(* Logix 5000 project; controller FV vendor 1 type 14 code 217 rev 31.11; software revision 31.00; part 39 of 63 *)
(* tags used below, declared in another part *)
   FV_FV10C : PlantItem;   // FV10C
   FV_FV10C_RawOutput : ALIAS FOR Remote_IO:2:O.Data.2;   // FV_FV10C FV 10 cone cooling valve
   FV_FV10J : PlantItem;   // FV10J
   FV_FV10J_RawOutput : ALIAS FOR Remote_IO:2:O.Data.3;   // FV_FV10J FV 10 jacket cooling valve
   FV_FV11C : PlantItem;   // FV11C
   FV_FV11C_RawOutput : ALIAS FOR Remote_IO:2:O.Data.4;   // FV_FV11C FV 11 cone cooling valve
   FV_FV11J : PlantItem;   // FV11J
   FV_FV11J_RawOutput : ALIAS FOR Remote_IO:2:O.Data.5;   // FV_FV11J FV 11 jacket cooling valve
   FV_FV12C : PlantItem;   // FV12C
   FV_FV12C_RawOutput : ALIAS FOR Remote_IO:2:O.Data.6;   // FV_FV12C FV 12 cone cooling valve
   FV_FV12J : PlantItem;   // FV12J
   FV_FV12J_RawOutput : ALIAS FOR Remote_IO:2:O.Data.7;   // FV_FV12J FV 12 jacket cooling valve
   FV_FV13C : PlantItem;   // FV13C
   FV_FV13C_RawOutput : ALIAS FOR Remote_IO:2:O.Data.8;   // FV_FV13C FV 13 cone cooling valve
   FV_FV13J : PlantItem;   // FV13J
   FV_FV13J_RawOutput : ALIAS FOR Remote_IO:2:O.Data.9;   // FV_FV13J FV 13 jacket cooling valve
   FV_FV14C : PlantItem;   // FV14C
   FV_FV14C_RawOutput : ALIAS FOR Remote_IO:2:O.Data.10;   // FV_FV14C FV 14 cone cooling valve
   FV_FV14J : PlantItem;   // FV14J
   FV_FV14J_RawOutput : ALIAS FOR Remote_IO:2:O.Data.11;   // FV_FV14J FV 14 jacket cooling valve
   FV_FV15C : PlantItem;   // FV15C
   FV_FV15C_RawOutput : ALIAS FOR Remote_IO:2:O.Data.12;   // FV_FV15C FV 15 cone cooling valve
   FV_FV15J : PlantItem;   // FV15J
   FV_FV15J_RawOutput : ALIAS FOR Remote_IO:2:O.Data.13;   // FV_FV15J FV 15 jacket cooling valve
   FV_FV16C : PlantItem;   // FV16C
   FV_FV16C_RawOutput : ALIAS FOR Remote_IO:2:O.Data.14;   // FV_FV16C FV 16 cone cooling valve
   FV_FV16J : PlantItem;   // FV16J
   FV_FV16J_RawOutput : ALIAS FOR Remote_IO:2:O.Data.15;   // FV_FV16J FV 16 jacket cooling valve
   FV_FV17C : PlantItem;   // FV17C
   FV_FV17C_RawOutput : ALIAS FOR Remote_IO:3:O.Data.0;   // FV_FV17C FV 17 cone cooling valve
   FV_FV17J : PlantItem;   // FV17J
   FV_FV17J_RawOutput : ALIAS FOR Remote_IO:3:O.Data.1;   // FV_FV17J FV 17 jacket cooling valve
   FV_FV18C : PlantItem;   // FV18C
   FV_FV18C_RawOutput : ALIAS FOR Remote_IO:3:O.Data.2;   // FV_FV18C FV 18 cone cooling valve
   FV_FV18J : PlantItem;   // FV18J
   FV_FV18J_RawOutput : ALIAS FOR Remote_IO:3:O.Data.3;   // FV_FV18J FV 18 jacket cooling valve
   FV_FV19C : PlantItem;   // FV19C
   FV_FV19C_RawOutput : ALIAS FOR Remote_IO:3:O.Data.4;   // FV_FV19C FV 19 cone cooling valve
   FV_FV19J : PlantItem;   // FV19J
   FV_FV19J_RawOutput : ALIAS FOR Remote_IO:3:O.Data.5;   // FV_FV19J FV 19 jacket cooling valve
   FV_FV1C : PlantItem;   // FV1C
   FV_FV1C_RawOutput : ALIAS FOR Remote_IO:1:O.Data.0;   // FV_FV1C FV 1 cone cooling valve
   FV_FV1J : PlantItem;   // FV1J
   FV_FV1J_RawOutput : ALIAS FOR Remote_IO:1:O.Data.1;   // FV_FV1J FV 1 jacket cooling valve
   FV_FV20C : PlantItem;   // FV20C
   FV_FV20C_RawOutput : ALIAS FOR Remote_IO:3:O.Data.6;   // FV_FV20C FV 20 cone cooling valve
   FV_FV20J : PlantItem;   // FV20J
   FV_FV20J_RawOutput : ALIAS FOR Remote_IO:3:O.Data.7;   // FV_FV20J FV 20 jacket cooling valve
   FV_FV21C : PlantItem;   // FV21C
   FV_FV21C_RawOutput : ALIAS FOR Remote_IO:3:O.Data.8;   // FV_FV21C FV 21 cone cooling valve
   FV_FV21J : PlantItem;   // FV21J
   FV_FV21J_RawOutput : ALIAS FOR Remote_IO:3:O.Data.9;   // FV_FV21J FV 21 jacket cooling valve
   FV_FV22C : PlantItem;   // FV22C
   FV_FV22C_RawOutput : ALIAS FOR Remote_IO:3:O.Data.10;   // FV_FV22C FV 22 cone cooling valve
   FV_FV22J : PlantItem;   // FV22J
   FV_FV22J_RawOutput : ALIAS FOR Remote_IO:3:O.Data.11;   // FV_FV22J FV 22 jacket cooling valve
   FV_FV23C : PlantItem;   // FV23C
   FV_FV23C_RawOutput : ALIAS FOR Remote_IO:3:O.Data.12;   // FV_FV23C FV 23 cone cooling valve
   FV_FV23J : PlantItem;   // FV23J
   FV_FV23J_RawOutput : ALIAS FOR Remote_IO:3:O.Data.13;   // FV_FV23J FV 23 jacket cooling valve
   FV_FV24C : PlantItem;   // FV24C
   FV_FV24C_RawOutput : ALIAS FOR Remote_IO:3:O.Data.14;   // FV_FV24C FV 24 cone cooling valve
   FV_FV24J : PlantItem;   // FV24J
   FV_FV24J_RawOutput : ALIAS FOR Remote_IO:3:O.Data.15;   // FV_FV24J FV 24 jacket cooling valve
   FV_FV2C : PlantItem;   // FV2C
   FV_FV2C_RawOutput : ALIAS FOR Remote_IO:1:O.Data.2;   // FV_FV2C FV 2 cone cooling valve
   FV_FV2J : PlantItem;   // FV2J
   FV_FV2J_RawOutput : ALIAS FOR Remote_IO:1:O.Data.3;   // FV_FV2J FV 2 jacket cooling valve
   FV_FV3C : PlantItem;   // FV3C
   FV_FV3C_RawOutput : ALIAS FOR Remote_IO:1:O.Data.4;   // FV_FV3C FV 3 cone cooling valve
   FV_FV3J : PlantItem;   // FV3J
   FV_FV3J_RawOutput : ALIAS FOR Remote_IO:1:O.Data.5;   // FV_FV3J FV 3 jacket cooling valve
   FV_FV4C : PlantItem;   // FV4C
   FV_FV4C_RawOutput : ALIAS FOR Remote_IO:1:O.Data.6;   // FV_FV4C FV 4 cone cooling valve
   FV_FV4J : PlantItem;   // FV4J
   FV_FV4J_RawOutput : ALIAS FOR Remote_IO:1:O.Data.7;   // FV_FV4J FV 4 jacket cooling valve
   FV_FV5C : PlantItem;   // FV5C
   FV_FV5C_RawOutput : ALIAS FOR Remote_IO:1:O.Data.8;   // FV_FV5C FV 5 cone cooling valve
   FV_FV5J : PlantItem;   // FV5J
   FV_FV5J_RawOutput : ALIAS FOR Remote_IO:1:O.Data.9;   // FV_FV5J FV 5 jacket cooling valve
   FV_FV6C : PlantItem;   // FV6C
   FV_FV6C_RawOutput : ALIAS FOR Remote_IO:1:O.Data.10;   // FV_FV6C FV 6 cone cooling valve
   FV_FV6J : PlantItem;   // FV6J
   FV_FV6J_RawOutput : ALIAS FOR Remote_IO:1:O.Data.11;   // FV_FV6J FV 6 jacket cooling valve
   FV_FV7C : PlantItem;   // FV7C
   FV_FV7C_RawOutput : ALIAS FOR Remote_IO:1:O.Data.12;   // FV_FV7C FV 7 cone cooling valve
   FV_FV7J : PlantItem;   // FV7J
   FV_FV7J_RawOutput : ALIAS FOR Remote_IO:1:O.Data.13;   // FV_FV7J FV 7 jacket cooling valve
   FV_FV8C : PlantItem;   // FV8C
   FV_FV8C_RawOutput : ALIAS FOR Remote_IO:1:O.Data.14;   // FV_FV8C FV 8 cone cooling valve
   FV_FV8J : PlantItem;   // FV8J
   FV_FV8J_RawOutput : ALIAS FOR Remote_IO:1:O.Data.15;   // FV_FV8J FV 8 jacket cooling valve
   FV_FV9C : PlantItem;   // FV9C
   FV_FV9C_RawOutput : ALIAS FOR Remote_IO:2:O.Data.0;   // FV_FV9C FV 9 cone cooling valve
   FV_FV9J : PlantItem;   // FV9J
   FV_FV9J_RawOutput : ALIAS FOR Remote_IO:2:O.Data.1;   // FV_FV9J FV 9 jacket cooling valve
(* FV_Common, continued *)

ROUTINE FV_Digital_Outputs   (* ladder *)
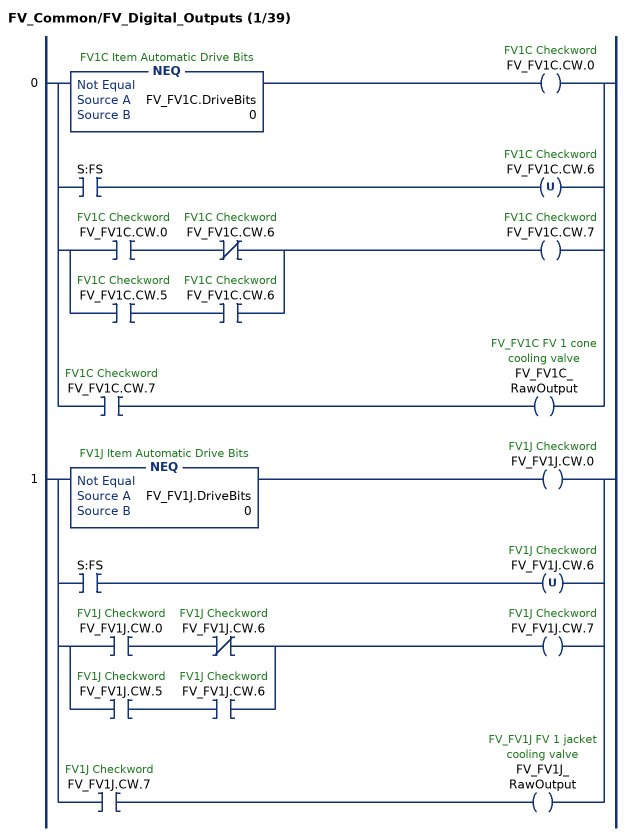
   0: [NEQ(FV_FV1C.DriveBits,0) OTE(FV_FV1C.CW.0) ,XIC(S:FS) OTU(FV_FV1C.CW.6) ,[XIC(FV_FV1C.CW.0) XIO(FV_FV1C.CW.6) ,XIC(FV_FV1C.CW.5) XIC(FV_FV1C.CW.6) ] OTE(FV_FV1C.CW.7) ,XIC(FV_FV1C.CW.7) OTE(FV_FV1C_RawOutput) ];
   1: [NEQ(FV_FV1J.DriveBits,0) OTE(FV_FV1J.CW.0) ,XIC(S:FS) OTU(FV_FV1J.CW.6) ,[XIC(FV_FV1J.CW.0) XIO(FV_FV1J.CW.6) ,XIC(FV_FV1J.CW.5) XIC(FV_FV1J.CW.6) ] OTE(FV_FV1J.CW.7) ,XIC(FV_FV1J.CW.7) OTE(FV_FV1J_RawOutput) ];
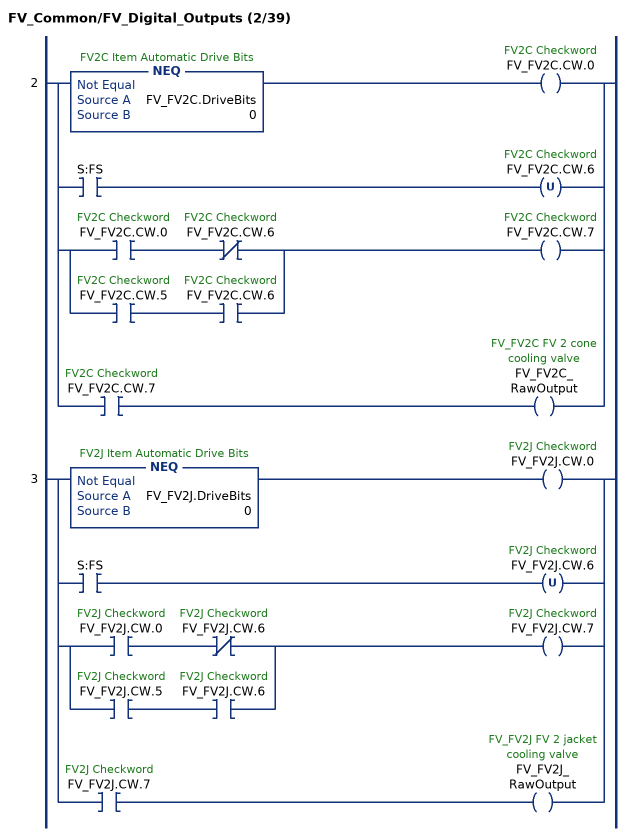
   2: [NEQ(FV_FV2C.DriveBits,0) OTE(FV_FV2C.CW.0) ,XIC(S:FS) OTU(FV_FV2C.CW.6) ,[XIC(FV_FV2C.CW.0) XIO(FV_FV2C.CW.6) ,XIC(FV_FV2C.CW.5) XIC(FV_FV2C.CW.6) ] OTE(FV_FV2C.CW.7) ,XIC(FV_FV2C.CW.7) OTE(FV_FV2C_RawOutput) ];
   3: [NEQ(FV_FV2J.DriveBits,0) OTE(FV_FV2J.CW.0) ,XIC(S:FS) OTU(FV_FV2J.CW.6) ,[XIC(FV_FV2J.CW.0) XIO(FV_FV2J.CW.6) ,XIC(FV_FV2J.CW.5) XIC(FV_FV2J.CW.6) ] OTE(FV_FV2J.CW.7) ,XIC(FV_FV2J.CW.7) OTE(FV_FV2J_RawOutput) ];
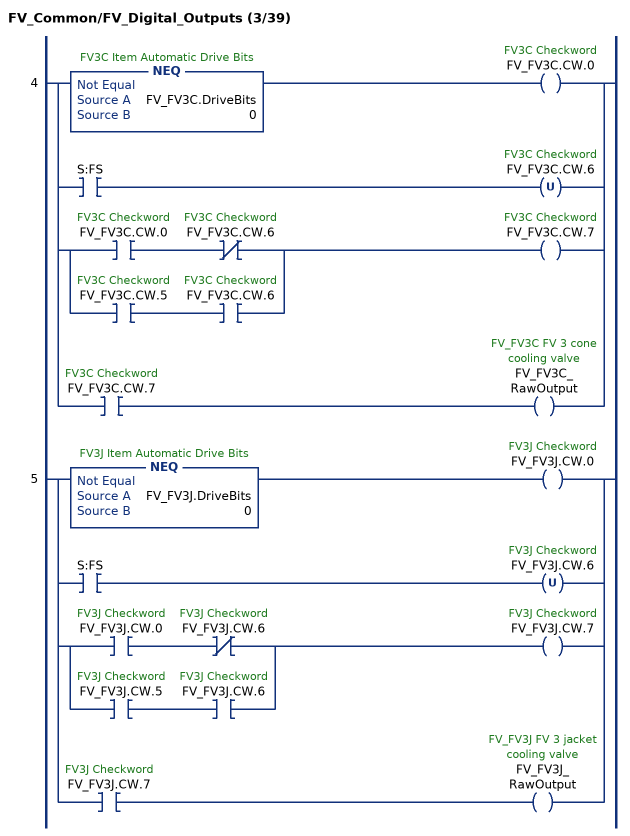
   4: [NEQ(FV_FV3C.DriveBits,0) OTE(FV_FV3C.CW.0) ,XIC(S:FS) OTU(FV_FV3C.CW.6) ,[XIC(FV_FV3C.CW.0) XIO(FV_FV3C.CW.6) ,XIC(FV_FV3C.CW.5) XIC(FV_FV3C.CW.6) ] OTE(FV_FV3C.CW.7) ,XIC(FV_FV3C.CW.7) OTE(FV_FV3C_RawOutput) ];
   5: [NEQ(FV_FV3J.DriveBits,0) OTE(FV_FV3J.CW.0) ,XIC(S:FS) OTU(FV_FV3J.CW.6) ,[XIC(FV_FV3J.CW.0) XIO(FV_FV3J.CW.6) ,XIC(FV_FV3J.CW.5) XIC(FV_FV3J.CW.6) ] OTE(FV_FV3J.CW.7) ,XIC(FV_FV3J.CW.7) OTE(FV_FV3J_RawOutput) ];
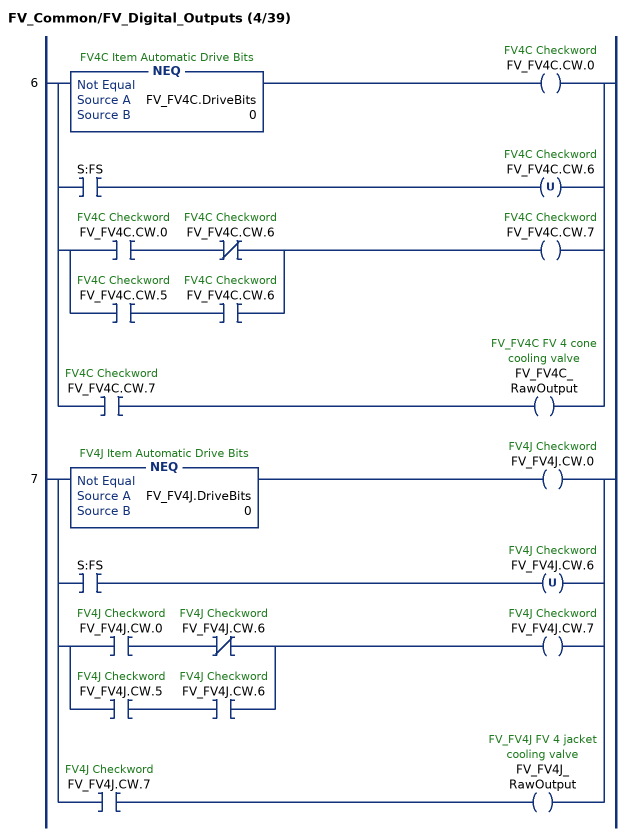
   6: [NEQ(FV_FV4C.DriveBits,0) OTE(FV_FV4C.CW.0) ,XIC(S:FS) OTU(FV_FV4C.CW.6) ,[XIC(FV_FV4C.CW.0) XIO(FV_FV4C.CW.6) ,XIC(FV_FV4C.CW.5) XIC(FV_FV4C.CW.6) ] OTE(FV_FV4C.CW.7) ,XIC(FV_FV4C.CW.7) OTE(FV_FV4C_RawOutput) ];
   7: [NEQ(FV_FV4J.DriveBits,0) OTE(FV_FV4J.CW.0) ,XIC(S:FS) OTU(FV_FV4J.CW.6) ,[XIC(FV_FV4J.CW.0) XIO(FV_FV4J.CW.6) ,XIC(FV_FV4J.CW.5) XIC(FV_FV4J.CW.6) ] OTE(FV_FV4J.CW.7) ,XIC(FV_FV4J.CW.7) OTE(FV_FV4J_RawOutput) ];
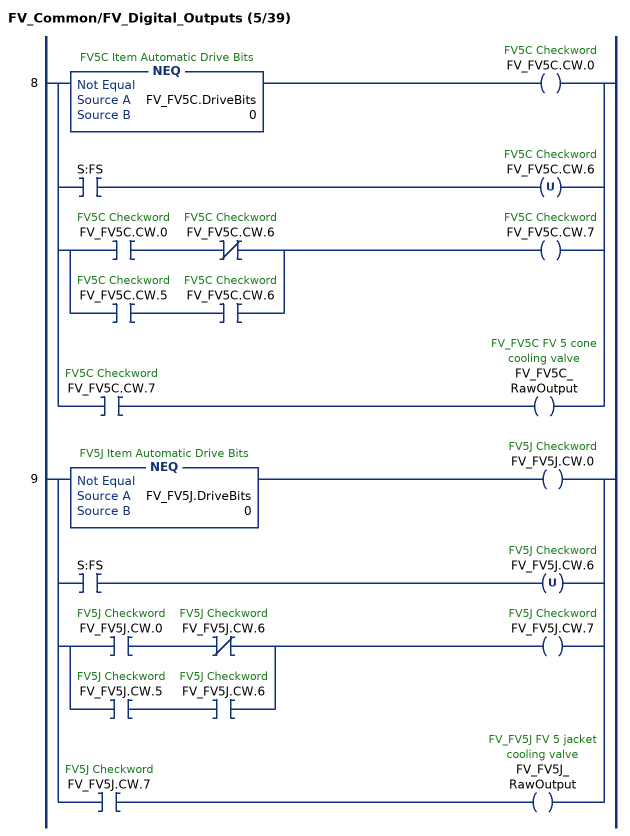
   8: [NEQ(FV_FV5C.DriveBits,0) OTE(FV_FV5C.CW.0) ,XIC(S:FS) OTU(FV_FV5C.CW.6) ,[XIC(FV_FV5C.CW.0) XIO(FV_FV5C.CW.6) ,XIC(FV_FV5C.CW.5) XIC(FV_FV5C.CW.6) ] OTE(FV_FV5C.CW.7) ,XIC(FV_FV5C.CW.7) OTE(FV_FV5C_RawOutput) ];
   9: [NEQ(FV_FV5J.DriveBits,0) OTE(FV_FV5J.CW.0) ,XIC(S:FS) OTU(FV_FV5J.CW.6) ,[XIC(FV_FV5J.CW.0) XIO(FV_FV5J.CW.6) ,XIC(FV_FV5J.CW.5) XIC(FV_FV5J.CW.6) ] OTE(FV_FV5J.CW.7) ,XIC(FV_FV5J.CW.7) OTE(FV_FV5J_RawOutput) ];
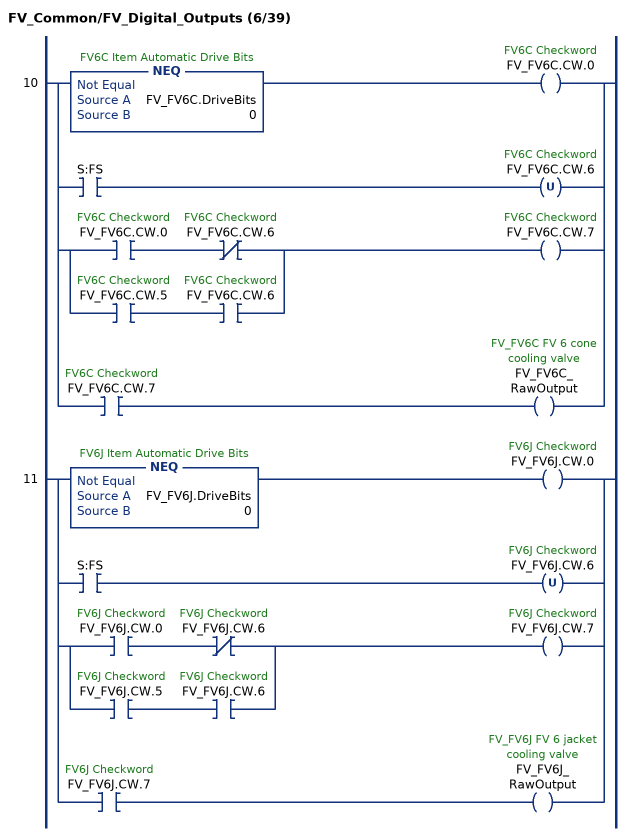
   10: [NEQ(FV_FV6C.DriveBits,0) OTE(FV_FV6C.CW.0) ,XIC(S:FS) OTU(FV_FV6C.CW.6) ,[XIC(FV_FV6C.CW.0) XIO(FV_FV6C.CW.6) ,XIC(FV_FV6C.CW.5) XIC(FV_FV6C.CW.6) ] OTE(FV_FV6C.CW.7) ,XIC(FV_FV6C.CW.7) OTE(FV_FV6C_RawOutput) ];
   11: [NEQ(FV_FV6J.DriveBits,0) OTE(FV_FV6J.CW.0) ,XIC(S:FS) OTU(FV_FV6J.CW.6) ,[XIC(FV_FV6J.CW.0) XIO(FV_FV6J.CW.6) ,XIC(FV_FV6J.CW.5) XIC(FV_FV6J.CW.6) ] OTE(FV_FV6J.CW.7) ,XIC(FV_FV6J.CW.7) OTE(FV_FV6J_RawOutput) ];
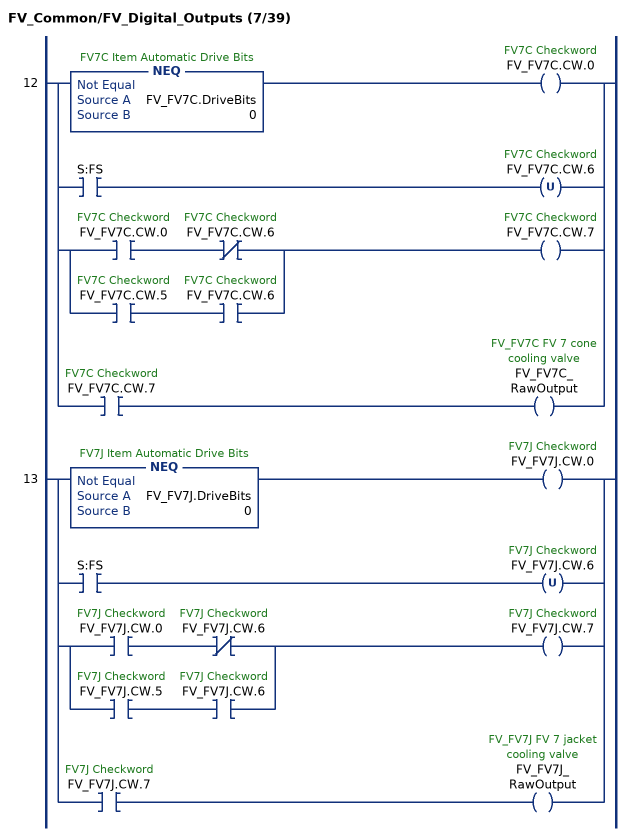
   12: [NEQ(FV_FV7C.DriveBits,0) OTE(FV_FV7C.CW.0) ,XIC(S:FS) OTU(FV_FV7C.CW.6) ,[XIC(FV_FV7C.CW.0) XIO(FV_FV7C.CW.6) ,XIC(FV_FV7C.CW.5) XIC(FV_FV7C.CW.6) ] OTE(FV_FV7C.CW.7) ,XIC(FV_FV7C.CW.7) OTE(FV_FV7C_RawOutput) ];
   13: [NEQ(FV_FV7J.DriveBits,0) OTE(FV_FV7J.CW.0) ,XIC(S:FS) OTU(FV_FV7J.CW.6) ,[XIC(FV_FV7J.CW.0) XIO(FV_FV7J.CW.6) ,XIC(FV_FV7J.CW.5) XIC(FV_FV7J.CW.6) ] OTE(FV_FV7J.CW.7) ,XIC(FV_FV7J.CW.7) OTE(FV_FV7J_RawOutput) ];
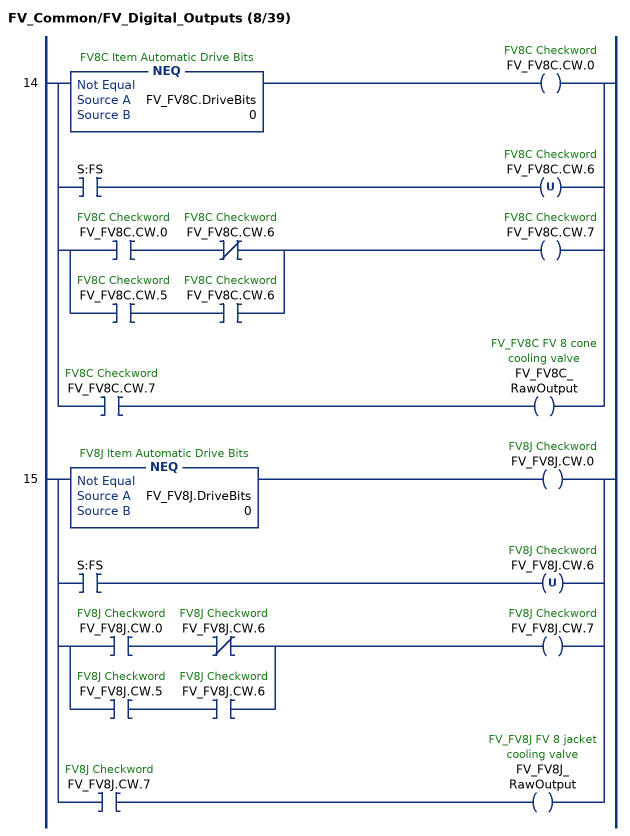
   14: [NEQ(FV_FV8C.DriveBits,0) OTE(FV_FV8C.CW.0) ,XIC(S:FS) OTU(FV_FV8C.CW.6) ,[XIC(FV_FV8C.CW.0) XIO(FV_FV8C.CW.6) ,XIC(FV_FV8C.CW.5) XIC(FV_FV8C.CW.6) ] OTE(FV_FV8C.CW.7) ,XIC(FV_FV8C.CW.7) OTE(FV_FV8C_RawOutput) ];
   15: [NEQ(FV_FV8J.DriveBits,0) OTE(FV_FV8J.CW.0) ,XIC(S:FS) OTU(FV_FV8J.CW.6) ,[XIC(FV_FV8J.CW.0) XIO(FV_FV8J.CW.6) ,XIC(FV_FV8J.CW.5) XIC(FV_FV8J.CW.6) ] OTE(FV_FV8J.CW.7) ,XIC(FV_FV8J.CW.7) OTE(FV_FV8J_RawOutput) ];
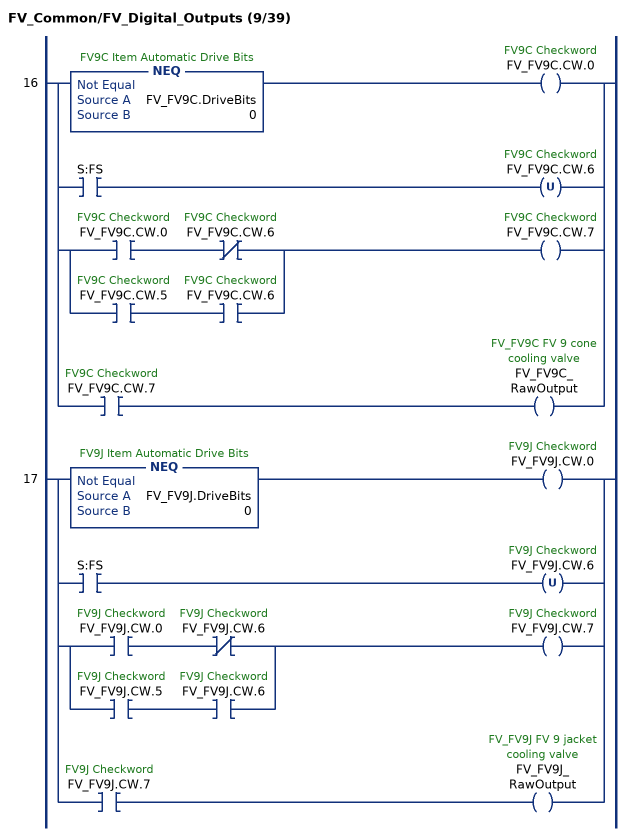
   16: [NEQ(FV_FV9C.DriveBits,0) OTE(FV_FV9C.CW.0) ,XIC(S:FS) OTU(FV_FV9C.CW.6) ,[XIC(FV_FV9C.CW.0) XIO(FV_FV9C.CW.6) ,XIC(FV_FV9C.CW.5) XIC(FV_FV9C.CW.6) ] OTE(FV_FV9C.CW.7) ,XIC(FV_FV9C.CW.7) OTE(FV_FV9C_RawOutput) ];
   17: [NEQ(FV_FV9J.DriveBits,0) OTE(FV_FV9J.CW.0) ,XIC(S:FS) OTU(FV_FV9J.CW.6) ,[XIC(FV_FV9J.CW.0) XIO(FV_FV9J.CW.6) ,XIC(FV_FV9J.CW.5) XIC(FV_FV9J.CW.6) ] OTE(FV_FV9J.CW.7) ,XIC(FV_FV9J.CW.7) OTE(FV_FV9J_RawOutput) ];
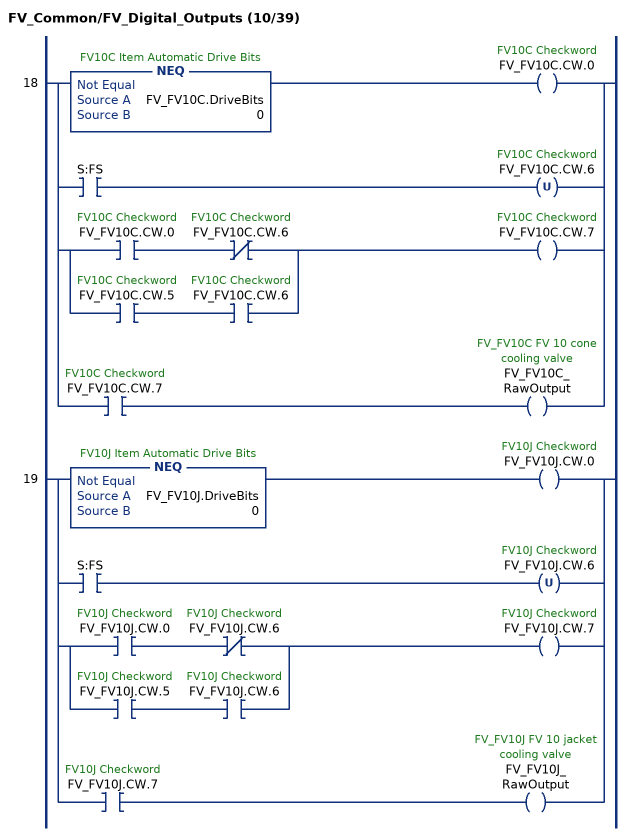
   18: [NEQ(FV_FV10C.DriveBits,0) OTE(FV_FV10C.CW.0) ,XIC(S:FS) OTU(FV_FV10C.CW.6) ,[XIC(FV_FV10C.CW.0) XIO(FV_FV10C.CW.6) ,XIC(FV_FV10C.CW.5) XIC(FV_FV10C.CW.6) ] OTE(FV_FV10C.CW.7) ,XIC(FV_FV10C.CW.7) OTE(FV_FV10C_RawOutput) ];
   19: [NEQ(FV_FV10J.DriveBits,0) OTE(FV_FV10J.CW.0) ,XIC(S:FS) OTU(FV_FV10J.CW.6) ,[XIC(FV_FV10J.CW.0) XIO(FV_FV10J.CW.6) ,XIC(FV_FV10J.CW.5) XIC(FV_FV10J.CW.6) ] OTE(FV_FV10J.CW.7) ,XIC(FV_FV10J.CW.7) OTE(FV_FV10J_RawOutput) ];
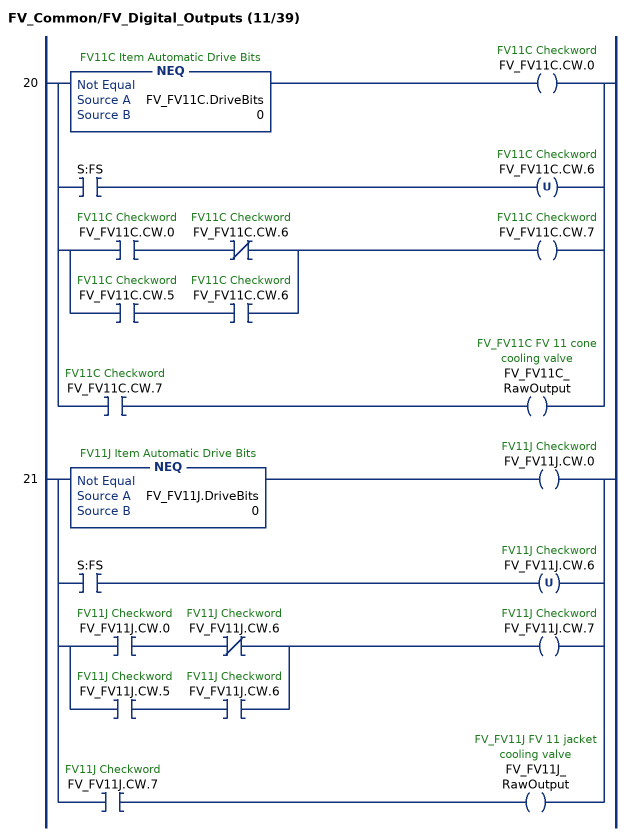
   20: [NEQ(FV_FV11C.DriveBits,0) OTE(FV_FV11C.CW.0) ,XIC(S:FS) OTU(FV_FV11C.CW.6) ,[XIC(FV_FV11C.CW.0) XIO(FV_FV11C.CW.6) ,XIC(FV_FV11C.CW.5) XIC(FV_FV11C.CW.6) ] OTE(FV_FV11C.CW.7) ,XIC(FV_FV11C.CW.7) OTE(FV_FV11C_RawOutput) ];
   21: [NEQ(FV_FV11J.DriveBits,0) OTE(FV_FV11J.CW.0) ,XIC(S:FS) OTU(FV_FV11J.CW.6) ,[XIC(FV_FV11J.CW.0) XIO(FV_FV11J.CW.6) ,XIC(FV_FV11J.CW.5) XIC(FV_FV11J.CW.6) ] OTE(FV_FV11J.CW.7) ,XIC(FV_FV11J.CW.7) OTE(FV_FV11J_RawOutput) ];
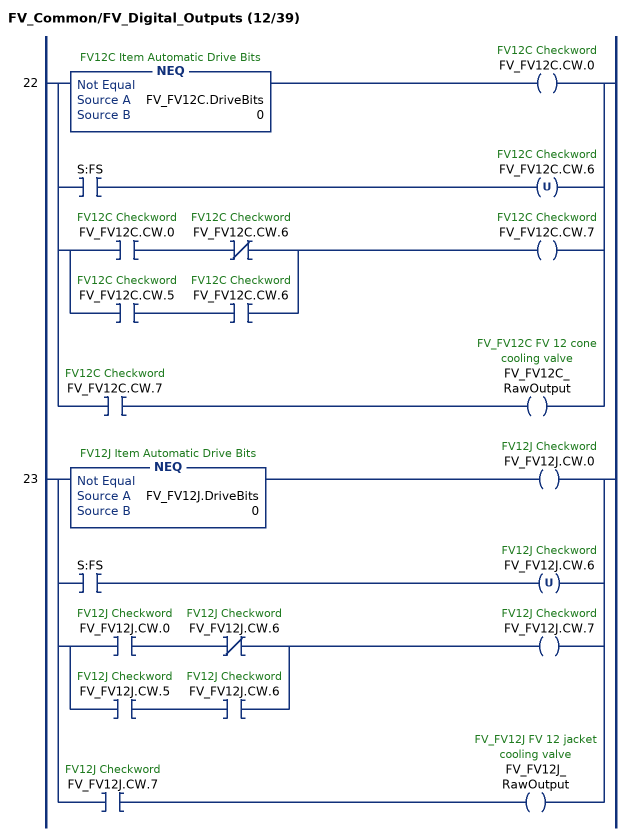
   22: [NEQ(FV_FV12C.DriveBits,0) OTE(FV_FV12C.CW.0) ,XIC(S:FS) OTU(FV_FV12C.CW.6) ,[XIC(FV_FV12C.CW.0) XIO(FV_FV12C.CW.6) ,XIC(FV_FV12C.CW.5) XIC(FV_FV12C.CW.6) ] OTE(FV_FV12C.CW.7) ,XIC(FV_FV12C.CW.7) OTE(FV_FV12C_RawOutput) ];
   23: [NEQ(FV_FV12J.DriveBits,0) OTE(FV_FV12J.CW.0) ,XIC(S:FS) OTU(FV_FV12J.CW.6) ,[XIC(FV_FV12J.CW.0) XIO(FV_FV12J.CW.6) ,XIC(FV_FV12J.CW.5) XIC(FV_FV12J.CW.6) ] OTE(FV_FV12J.CW.7) ,XIC(FV_FV12J.CW.7) OTE(FV_FV12J_RawOutput) ];
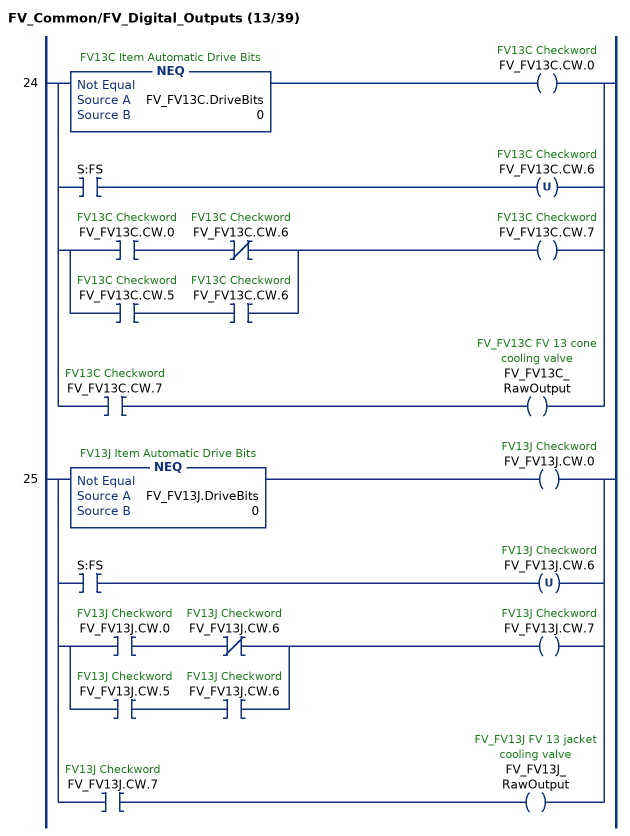
   24: [NEQ(FV_FV13C.DriveBits,0) OTE(FV_FV13C.CW.0) ,XIC(S:FS) OTU(FV_FV13C.CW.6) ,[XIC(FV_FV13C.CW.0) XIO(FV_FV13C.CW.6) ,XIC(FV_FV13C.CW.5) XIC(FV_FV13C.CW.6) ] OTE(FV_FV13C.CW.7) ,XIC(FV_FV13C.CW.7) OTE(FV_FV13C_RawOutput) ];
   25: [NEQ(FV_FV13J.DriveBits,0) OTE(FV_FV13J.CW.0) ,XIC(S:FS) OTU(FV_FV13J.CW.6) ,[XIC(FV_FV13J.CW.0) XIO(FV_FV13J.CW.6) ,XIC(FV_FV13J.CW.5) XIC(FV_FV13J.CW.6) ] OTE(FV_FV13J.CW.7) ,XIC(FV_FV13J.CW.7) OTE(FV_FV13J_RawOutput) ];
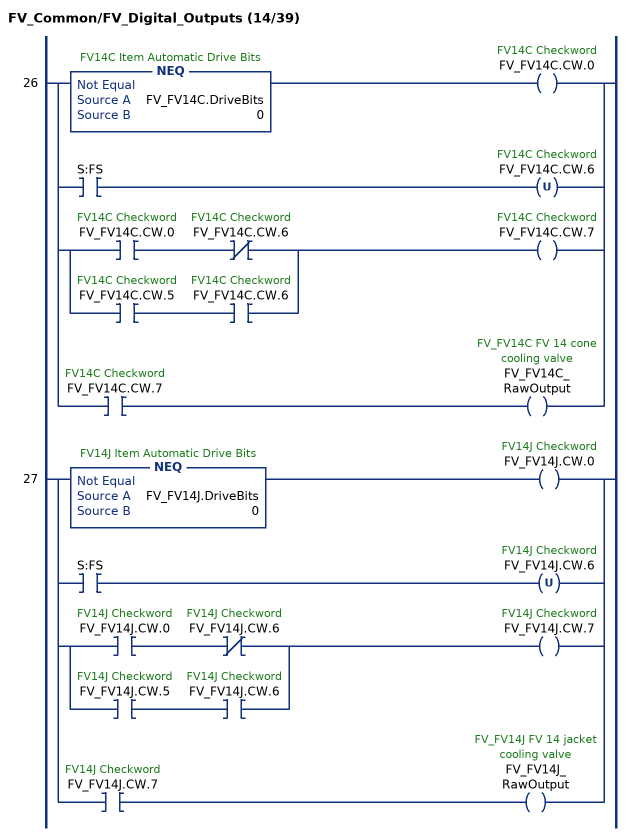
   26: [NEQ(FV_FV14C.DriveBits,0) OTE(FV_FV14C.CW.0) ,XIC(S:FS) OTU(FV_FV14C.CW.6) ,[XIC(FV_FV14C.CW.0) XIO(FV_FV14C.CW.6) ,XIC(FV_FV14C.CW.5) XIC(FV_FV14C.CW.6) ] OTE(FV_FV14C.CW.7) ,XIC(FV_FV14C.CW.7) OTE(FV_FV14C_RawOutput) ];
   27: [NEQ(FV_FV14J.DriveBits,0) OTE(FV_FV14J.CW.0) ,XIC(S:FS) OTU(FV_FV14J.CW.6) ,[XIC(FV_FV14J.CW.0) XIO(FV_FV14J.CW.6) ,XIC(FV_FV14J.CW.5) XIC(FV_FV14J.CW.6) ] OTE(FV_FV14J.CW.7) ,XIC(FV_FV14J.CW.7) OTE(FV_FV14J_RawOutput) ];
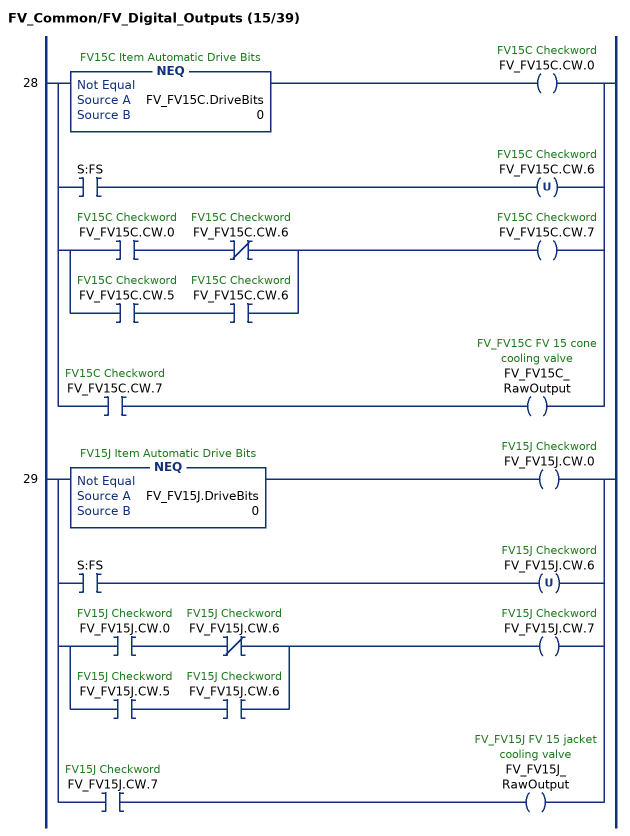
   28: [NEQ(FV_FV15C.DriveBits,0) OTE(FV_FV15C.CW.0) ,XIC(S:FS) OTU(FV_FV15C.CW.6) ,[XIC(FV_FV15C.CW.0) XIO(FV_FV15C.CW.6) ,XIC(FV_FV15C.CW.5) XIC(FV_FV15C.CW.6) ] OTE(FV_FV15C.CW.7) ,XIC(FV_FV15C.CW.7) OTE(FV_FV15C_RawOutput) ];
   29: [NEQ(FV_FV15J.DriveBits,0) OTE(FV_FV15J.CW.0) ,XIC(S:FS) OTU(FV_FV15J.CW.6) ,[XIC(FV_FV15J.CW.0) XIO(FV_FV15J.CW.6) ,XIC(FV_FV15J.CW.5) XIC(FV_FV15J.CW.6) ] OTE(FV_FV15J.CW.7) ,XIC(FV_FV15J.CW.7) OTE(FV_FV15J_RawOutput) ];
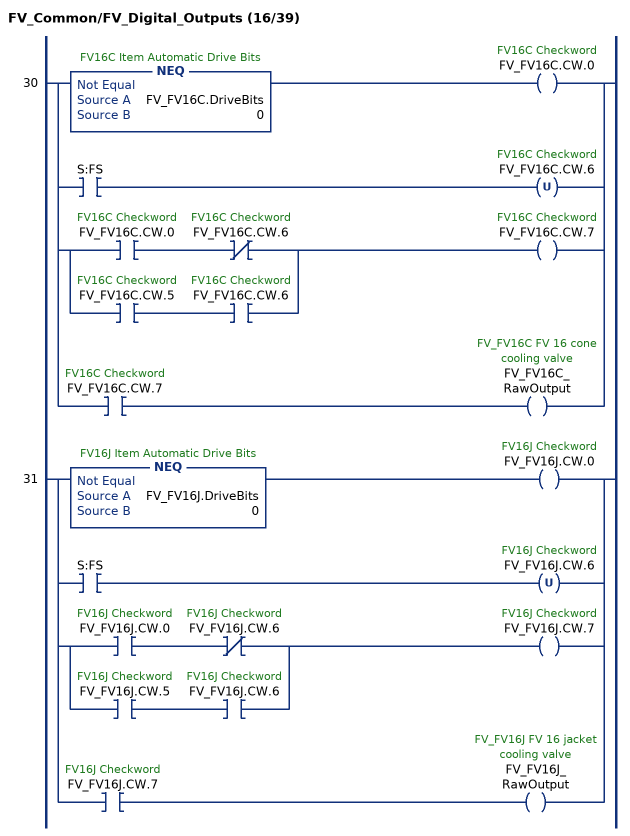
   30: [NEQ(FV_FV16C.DriveBits,0) OTE(FV_FV16C.CW.0) ,XIC(S:FS) OTU(FV_FV16C.CW.6) ,[XIC(FV_FV16C.CW.0) XIO(FV_FV16C.CW.6) ,XIC(FV_FV16C.CW.5) XIC(FV_FV16C.CW.6) ] OTE(FV_FV16C.CW.7) ,XIC(FV_FV16C.CW.7) OTE(FV_FV16C_RawOutput) ];
   31: [NEQ(FV_FV16J.DriveBits,0) OTE(FV_FV16J.CW.0) ,XIC(S:FS) OTU(FV_FV16J.CW.6) ,[XIC(FV_FV16J.CW.0) XIO(FV_FV16J.CW.6) ,XIC(FV_FV16J.CW.5) XIC(FV_FV16J.CW.6) ] OTE(FV_FV16J.CW.7) ,XIC(FV_FV16J.CW.7) OTE(FV_FV16J_RawOutput) ];
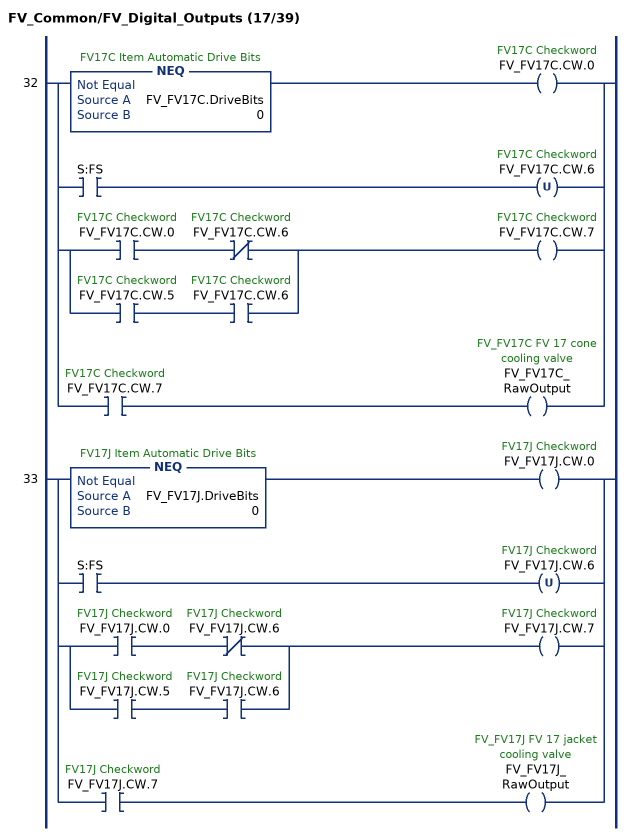
   32: [NEQ(FV_FV17C.DriveBits,0) OTE(FV_FV17C.CW.0) ,XIC(S:FS) OTU(FV_FV17C.CW.6) ,[XIC(FV_FV17C.CW.0) XIO(FV_FV17C.CW.6) ,XIC(FV_FV17C.CW.5) XIC(FV_FV17C.CW.6) ] OTE(FV_FV17C.CW.7) ,XIC(FV_FV17C.CW.7) OTE(FV_FV17C_RawOutput) ];
   33: [NEQ(FV_FV17J.DriveBits,0) OTE(FV_FV17J.CW.0) ,XIC(S:FS) OTU(FV_FV17J.CW.6) ,[XIC(FV_FV17J.CW.0) XIO(FV_FV17J.CW.6) ,XIC(FV_FV17J.CW.5) XIC(FV_FV17J.CW.6) ] OTE(FV_FV17J.CW.7) ,XIC(FV_FV17J.CW.7) OTE(FV_FV17J_RawOutput) ];
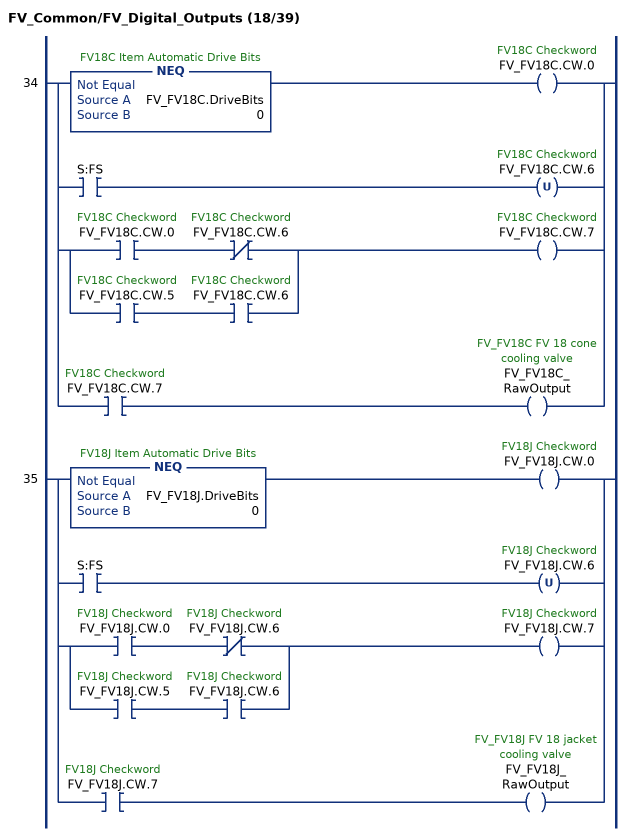
   34: [NEQ(FV_FV18C.DriveBits,0) OTE(FV_FV18C.CW.0) ,XIC(S:FS) OTU(FV_FV18C.CW.6) ,[XIC(FV_FV18C.CW.0) XIO(FV_FV18C.CW.6) ,XIC(FV_FV18C.CW.5) XIC(FV_FV18C.CW.6) ] OTE(FV_FV18C.CW.7) ,XIC(FV_FV18C.CW.7) OTE(FV_FV18C_RawOutput) ];
   35: [NEQ(FV_FV18J.DriveBits,0) OTE(FV_FV18J.CW.0) ,XIC(S:FS) OTU(FV_FV18J.CW.6) ,[XIC(FV_FV18J.CW.0) XIO(FV_FV18J.CW.6) ,XIC(FV_FV18J.CW.5) XIC(FV_FV18J.CW.6) ] OTE(FV_FV18J.CW.7) ,XIC(FV_FV18J.CW.7) OTE(FV_FV18J_RawOutput) ];
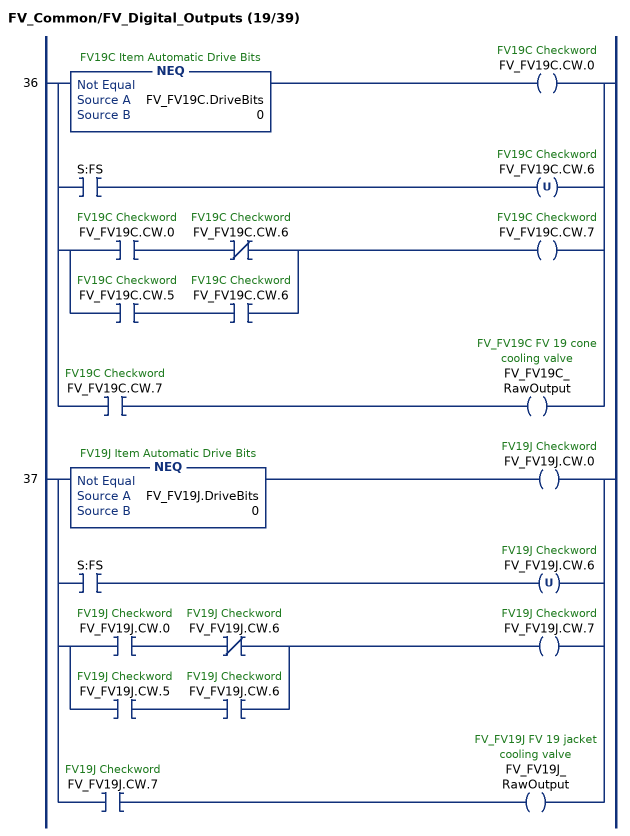
   36: [NEQ(FV_FV19C.DriveBits,0) OTE(FV_FV19C.CW.0) ,XIC(S:FS) OTU(FV_FV19C.CW.6) ,[XIC(FV_FV19C.CW.0) XIO(FV_FV19C.CW.6) ,XIC(FV_FV19C.CW.5) XIC(FV_FV19C.CW.6) ] OTE(FV_FV19C.CW.7) ,XIC(FV_FV19C.CW.7) OTE(FV_FV19C_RawOutput) ];
   37: [NEQ(FV_FV19J.DriveBits,0) OTE(FV_FV19J.CW.0) ,XIC(S:FS) OTU(FV_FV19J.CW.6) ,[XIC(FV_FV19J.CW.0) XIO(FV_FV19J.CW.6) ,XIC(FV_FV19J.CW.5) XIC(FV_FV19J.CW.6) ] OTE(FV_FV19J.CW.7) ,XIC(FV_FV19J.CW.7) OTE(FV_FV19J_RawOutput) ];
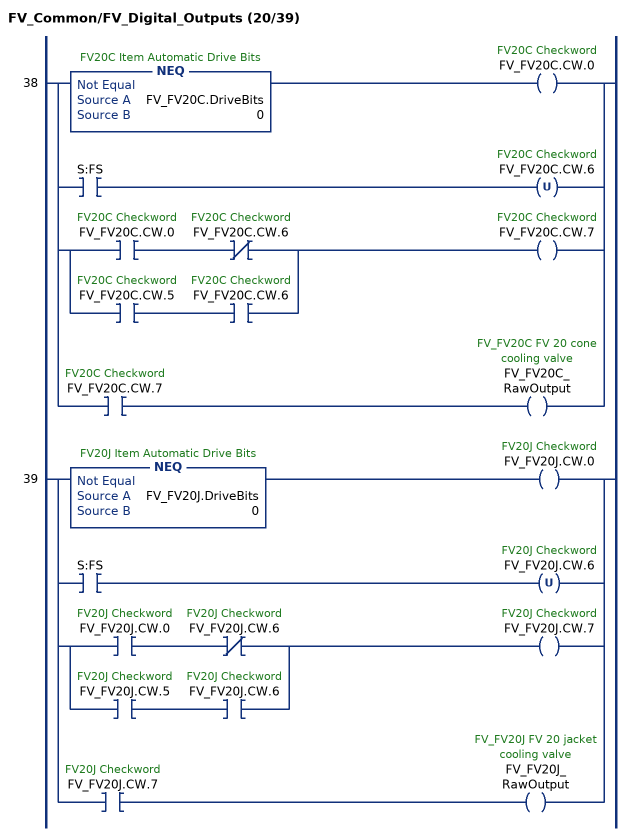
   38: [NEQ(FV_FV20C.DriveBits,0) OTE(FV_FV20C.CW.0) ,XIC(S:FS) OTU(FV_FV20C.CW.6) ,[XIC(FV_FV20C.CW.0) XIO(FV_FV20C.CW.6) ,XIC(FV_FV20C.CW.5) XIC(FV_FV20C.CW.6) ] OTE(FV_FV20C.CW.7) ,XIC(FV_FV20C.CW.7) OTE(FV_FV20C_RawOutput) ];
   39: [NEQ(FV_FV20J.DriveBits,0) OTE(FV_FV20J.CW.0) ,XIC(S:FS) OTU(FV_FV20J.CW.6) ,[XIC(FV_FV20J.CW.0) XIO(FV_FV20J.CW.6) ,XIC(FV_FV20J.CW.5) XIC(FV_FV20J.CW.6) ] OTE(FV_FV20J.CW.7) ,XIC(FV_FV20J.CW.7) OTE(FV_FV20J_RawOutput) ];
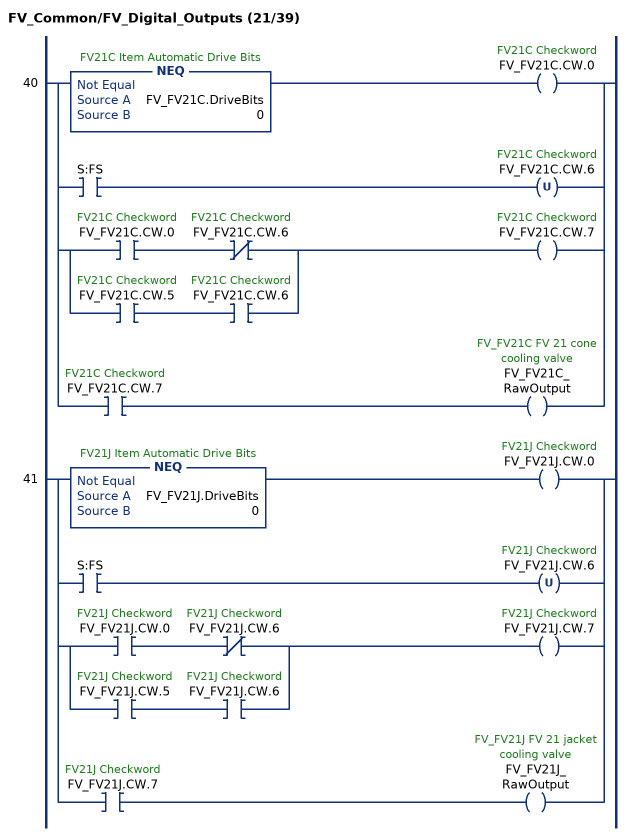
   40: [NEQ(FV_FV21C.DriveBits,0) OTE(FV_FV21C.CW.0) ,XIC(S:FS) OTU(FV_FV21C.CW.6) ,[XIC(FV_FV21C.CW.0) XIO(FV_FV21C.CW.6) ,XIC(FV_FV21C.CW.5) XIC(FV_FV21C.CW.6) ] OTE(FV_FV21C.CW.7) ,XIC(FV_FV21C.CW.7) OTE(FV_FV21C_RawOutput) ];
   41: [NEQ(FV_FV21J.DriveBits,0) OTE(FV_FV21J.CW.0) ,XIC(S:FS) OTU(FV_FV21J.CW.6) ,[XIC(FV_FV21J.CW.0) XIO(FV_FV21J.CW.6) ,XIC(FV_FV21J.CW.5) XIC(FV_FV21J.CW.6) ] OTE(FV_FV21J.CW.7) ,XIC(FV_FV21J.CW.7) OTE(FV_FV21J_RawOutput) ];
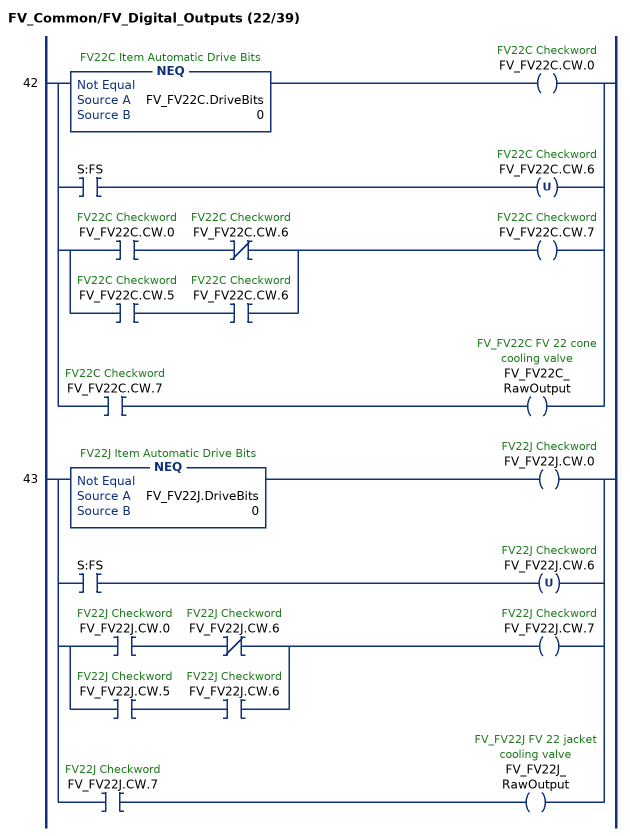
   42: [NEQ(FV_FV22C.DriveBits,0) OTE(FV_FV22C.CW.0) ,XIC(S:FS) OTU(FV_FV22C.CW.6) ,[XIC(FV_FV22C.CW.0) XIO(FV_FV22C.CW.6) ,XIC(FV_FV22C.CW.5) XIC(FV_FV22C.CW.6) ] OTE(FV_FV22C.CW.7) ,XIC(FV_FV22C.CW.7) OTE(FV_FV22C_RawOutput) ];
   43: [NEQ(FV_FV22J.DriveBits,0) OTE(FV_FV22J.CW.0) ,XIC(S:FS) OTU(FV_FV22J.CW.6) ,[XIC(FV_FV22J.CW.0) XIO(FV_FV22J.CW.6) ,XIC(FV_FV22J.CW.5) XIC(FV_FV22J.CW.6) ] OTE(FV_FV22J.CW.7) ,XIC(FV_FV22J.CW.7) OTE(FV_FV22J_RawOutput) ];
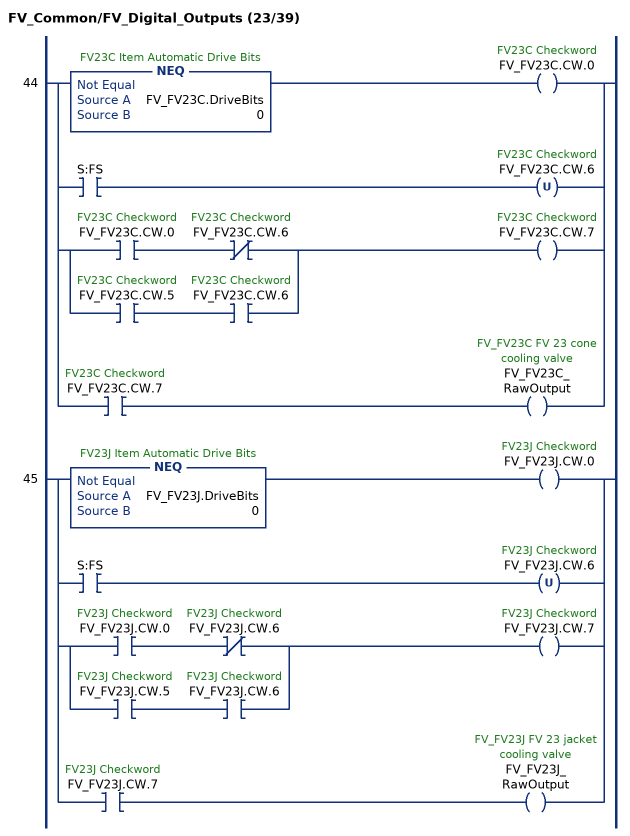
   44: [NEQ(FV_FV23C.DriveBits,0) OTE(FV_FV23C.CW.0) ,XIC(S:FS) OTU(FV_FV23C.CW.6) ,[XIC(FV_FV23C.CW.0) XIO(FV_FV23C.CW.6) ,XIC(FV_FV23C.CW.5) XIC(FV_FV23C.CW.6) ] OTE(FV_FV23C.CW.7) ,XIC(FV_FV23C.CW.7) OTE(FV_FV23C_RawOutput) ];
   45: [NEQ(FV_FV23J.DriveBits,0) OTE(FV_FV23J.CW.0) ,XIC(S:FS) OTU(FV_FV23J.CW.6) ,[XIC(FV_FV23J.CW.0) XIO(FV_FV23J.CW.6) ,XIC(FV_FV23J.CW.5) XIC(FV_FV23J.CW.6) ] OTE(FV_FV23J.CW.7) ,XIC(FV_FV23J.CW.7) OTE(FV_FV23J_RawOutput) ];
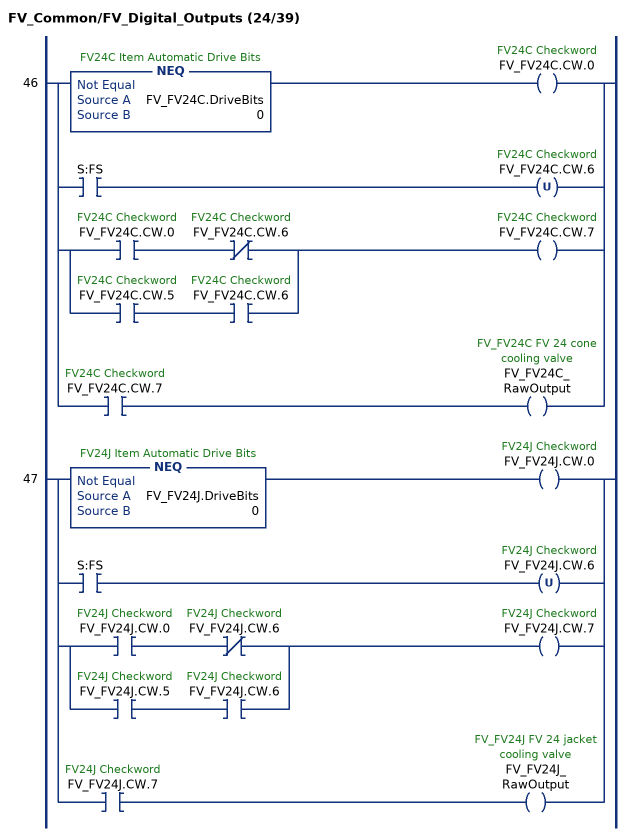
   46: [NEQ(FV_FV24C.DriveBits,0) OTE(FV_FV24C.CW.0) ,XIC(S:FS) OTU(FV_FV24C.CW.6) ,[XIC(FV_FV24C.CW.0) XIO(FV_FV24C.CW.6) ,XIC(FV_FV24C.CW.5) XIC(FV_FV24C.CW.6) ] OTE(FV_FV24C.CW.7) ,XIC(FV_FV24C.CW.7) OTE(FV_FV24C_RawOutput) ];
   47: [NEQ(FV_FV24J.DriveBits,0) OTE(FV_FV24J.CW.0) ,XIC(S:FS) OTU(FV_FV24J.CW.6) ,[XIC(FV_FV24J.CW.0) XIO(FV_FV24J.CW.6) ,XIC(FV_FV24J.CW.5) XIC(FV_FV24J.CW.6) ] OTE(FV_FV24J.CW.7) ,XIC(FV_FV24J.CW.7) OTE(FV_FV24J_RawOutput) ];
